// TIA Portal project "消毒机" (V15.1) (continued)
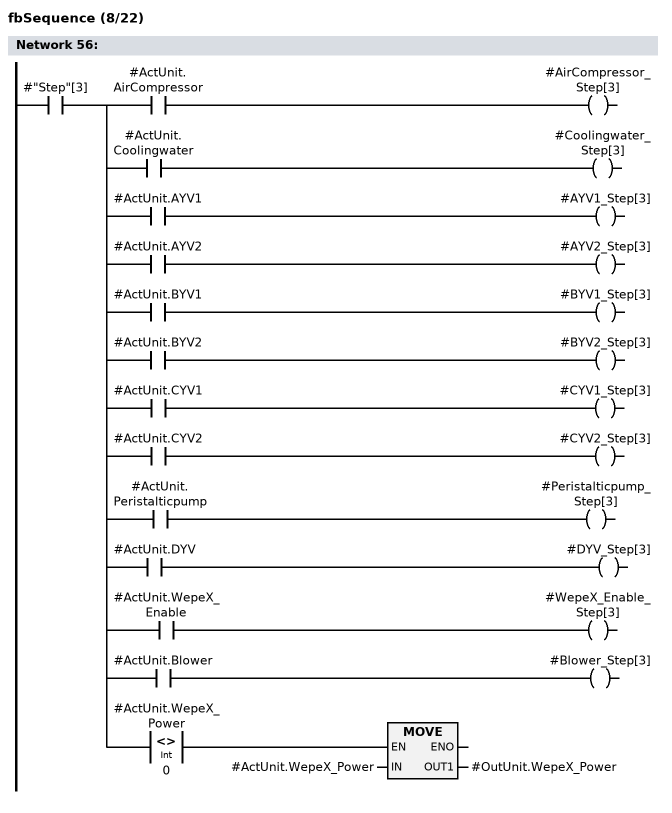
   RUNG wire#powerrail
      Contact( #"Step"[3] )
      wire#w1
      Contact( #ActUnit.AirCompressor )
      Coil( #AirCompressor_Step[3] )
   END_RUNG
   RUNG wire#w1
      Contact( #ActUnit.Coolingwater )
      Coil( #Coolingwater_Step[3] )
   END_RUNG
   RUNG wire#w1
      Contact( #ActUnit.AYV1 )
      Coil( #AYV1_Step[3] )
   END_RUNG
   RUNG wire#w1
      Contact( #ActUnit.AYV2 )
      Coil( #AYV2_Step[3] )
   END_RUNG
   RUNG wire#w1
      Contact( #ActUnit.BYV1 )
      Coil( #BYV1_Step[3] )
   END_RUNG
   RUNG wire#w1
      Contact( #ActUnit.BYV2 )
      Coil( #BYV2_Step[3] )
   END_RUNG
   RUNG wire#w1
      Contact( #ActUnit.CYV1 )
      Coil( #CYV1_Step[3] )
   END_RUNG
   RUNG wire#w1
      Contact( #ActUnit.CYV2 )
      Coil( #CYV2_Step[3] )
   END_RUNG
   RUNG wire#w1
      Contact( #ActUnit.Peristalticpump )
      Coil( #Peristalticpump_Step[3] )
   END_RUNG
   RUNG wire#w1
      Contact( #ActUnit.DYV )
      Coil( #DYV_Step[3] )
   END_RUNG
   RUNG wire#w1
      Contact( #ActUnit.WepeX_Enable )
      Coil( #WepeX_Enable_Step[3] )
   END_RUNG
   RUNG wire#w1
      Contact( #ActUnit.Blower )
      Coil( #Blower_Step[3] )
   END_RUNG
   RUNG wire#w1
      { S7_Templates := "SrcType := Int" } NE_Contact(in1 := #ActUnit.WepeX_Power, in2 := 0)
      Move(in := #ActUnit.WepeX_Power, out1 => #OutUnit.WepeX_Power)
   END_RUNG
   // the same network as SCL:
   #AirCompressor_Step[3] := #"Step"[3] AND #ActUnit.AirCompressor;
   #Coolingwater_Step[3] := #"Step"[3] AND #ActUnit.Coolingwater;
   #AYV1_Step[3] := #"Step"[3] AND #ActUnit.AYV1;
   #AYV2_Step[3] := #"Step"[3] AND #ActUnit.AYV2;
   #BYV1_Step[3] := #"Step"[3] AND #ActUnit.BYV1;
   #BYV2_Step[3] := #"Step"[3] AND #ActUnit.BYV2;
   #CYV1_Step[3] := #"Step"[3] AND #ActUnit.CYV1;
   #CYV2_Step[3] := #"Step"[3] AND #ActUnit.CYV2;
   #Peristalticpump_Step[3] := #"Step"[3] AND #ActUnit.Peristalticpump;
   #DYV_Step[3] := #"Step"[3] AND #ActUnit.DYV;
   #WepeX_Enable_Step[3] := #"Step"[3] AND #ActUnit.WepeX_Enable;
   #Blower_Step[3] := #"Step"[3] AND #ActUnit.Blower;
   IF #"Step"[3] AND (#ActUnit.WepeX_Power <> 0) THEN #OutUnit.WepeX_Power := #ActUnit.WepeX_Power; END_IF;
END_REGION

REGION Network 57
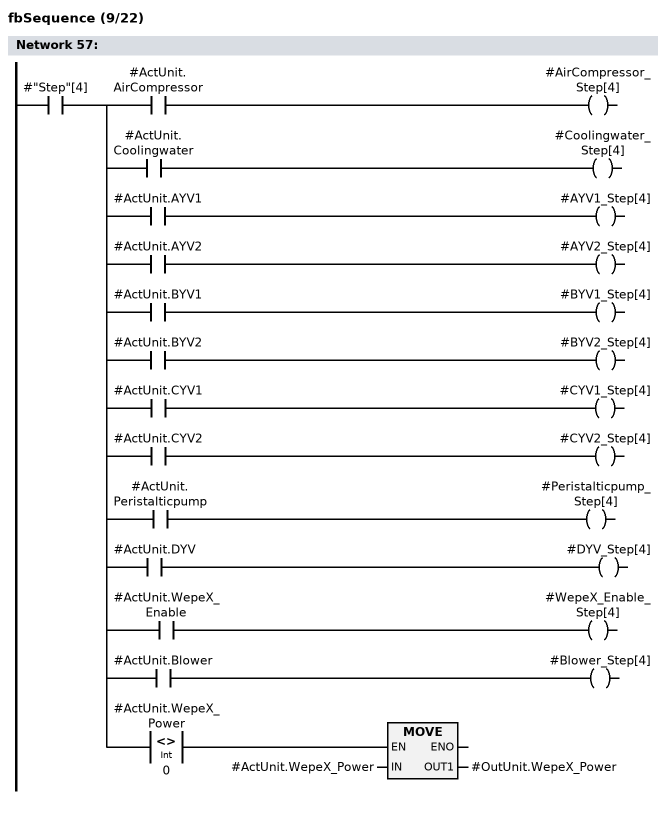
   RUNG wire#powerrail
      Contact( #"Step"[4] )
      wire#w1
      Contact( #ActUnit.AirCompressor )
      Coil( #AirCompressor_Step[4] )
   END_RUNG
   RUNG wire#w1
      Contact( #ActUnit.Coolingwater )
      Coil( #Coolingwater_Step[4] )
   END_RUNG
   RUNG wire#w1
      Contact( #ActUnit.AYV1 )
      Coil( #AYV1_Step[4] )
   END_RUNG
   RUNG wire#w1
      Contact( #ActUnit.AYV2 )
      Coil( #AYV2_Step[4] )
   END_RUNG
   RUNG wire#w1
      Contact( #ActUnit.BYV1 )
      Coil( #BYV1_Step[4] )
   END_RUNG
   RUNG wire#w1
      Contact( #ActUnit.BYV2 )
      Coil( #BYV2_Step[4] )
   END_RUNG
   RUNG wire#w1
      Contact( #ActUnit.CYV1 )
      Coil( #CYV1_Step[4] )
   END_RUNG
   RUNG wire#w1
      Contact( #ActUnit.CYV2 )
      Coil( #CYV2_Step[4] )
   END_RUNG
   RUNG wire#w1
      Contact( #ActUnit.Peristalticpump )
      Coil( #Peristalticpump_Step[4] )
   END_RUNG
   RUNG wire#w1
      Contact( #ActUnit.DYV )
      Coil( #DYV_Step[4] )
   END_RUNG
   RUNG wire#w1
      Contact( #ActUnit.WepeX_Enable )
      Coil( #WepeX_Enable_Step[4] )
   END_RUNG
   RUNG wire#w1
      Contact( #ActUnit.Blower )
      Coil( #Blower_Step[4] )
   END_RUNG
   RUNG wire#w1
      { S7_Templates := "SrcType := Int" } NE_Contact(in1 := #ActUnit.WepeX_Power, in2 := 0)
      Move(in := #ActUnit.WepeX_Power, out1 => #OutUnit.WepeX_Power)
   END_RUNG
   // the same network as SCL:
   #AirCompressor_Step[4] := #"Step"[4] AND #ActUnit.AirCompressor;
   #Coolingwater_Step[4] := #"Step"[4] AND #ActUnit.Coolingwater;
   #AYV1_Step[4] := #"Step"[4] AND #ActUnit.AYV1;
   #AYV2_Step[4] := #"Step"[4] AND #ActUnit.AYV2;
   #BYV1_Step[4] := #"Step"[4] AND #ActUnit.BYV1;
   #BYV2_Step[4] := #"Step"[4] AND #ActUnit.BYV2;
   #CYV1_Step[4] := #"Step"[4] AND #ActUnit.CYV1;
   #CYV2_Step[4] := #"Step"[4] AND #ActUnit.CYV2;
   #Peristalticpump_Step[4] := #"Step"[4] AND #ActUnit.Peristalticpump;
   #DYV_Step[4] := #"Step"[4] AND #ActUnit.DYV;
   #WepeX_Enable_Step[4] := #"Step"[4] AND #ActUnit.WepeX_Enable;
   #Blower_Step[4] := #"Step"[4] AND #ActUnit.Blower;
   IF #"Step"[4] AND (#ActUnit.WepeX_Power <> 0) THEN #OutUnit.WepeX_Power := #ActUnit.WepeX_Power; END_IF;
END_REGION

REGION Network 58
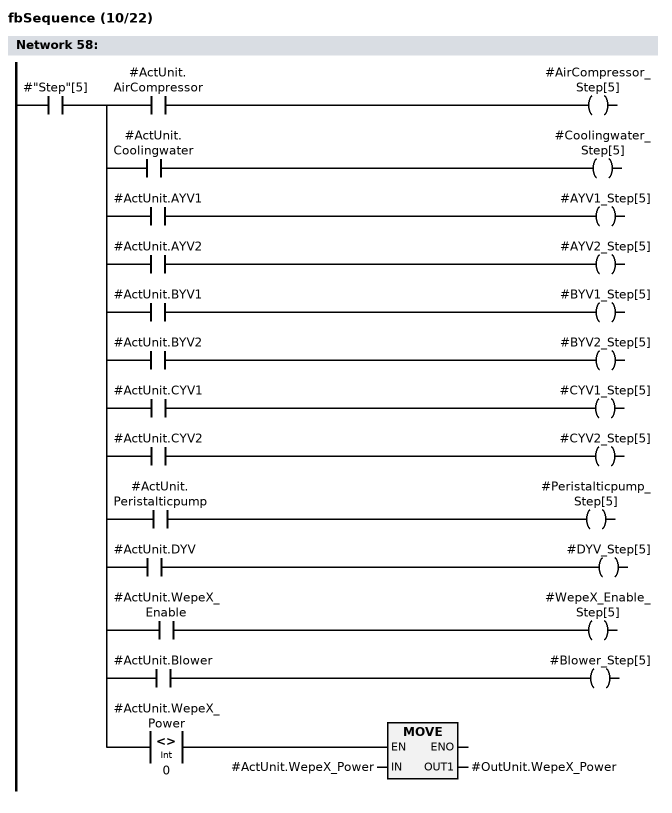
   RUNG wire#powerrail
      Contact( #"Step"[5] )
      wire#w1
      Contact( #ActUnit.AirCompressor )
      Coil( #AirCompressor_Step[5] )
   END_RUNG
   RUNG wire#w1
      Contact( #ActUnit.Coolingwater )
      Coil( #Coolingwater_Step[5] )
   END_RUNG
   RUNG wire#w1
      Contact( #ActUnit.AYV1 )
      Coil( #AYV1_Step[5] )
   END_RUNG
   RUNG wire#w1
      Contact( #ActUnit.AYV2 )
      Coil( #AYV2_Step[5] )
   END_RUNG
   RUNG wire#w1
      Contact( #ActUnit.BYV1 )
      Coil( #BYV1_Step[5] )
   END_RUNG
   RUNG wire#w1
      Contact( #ActUnit.BYV2 )
      Coil( #BYV2_Step[5] )
   END_RUNG
   RUNG wire#w1
      Contact( #ActUnit.CYV1 )
      Coil( #CYV1_Step[5] )
   END_RUNG
   RUNG wire#w1
      Contact( #ActUnit.CYV2 )
      Coil( #CYV2_Step[5] )
   END_RUNG
   RUNG wire#w1
      Contact( #ActUnit.Peristalticpump )
      Coil( #Peristalticpump_Step[5] )
   END_RUNG
   RUNG wire#w1
      Contact( #ActUnit.DYV )
      Coil( #DYV_Step[5] )
   END_RUNG
   RUNG wire#w1
      Contact( #ActUnit.WepeX_Enable )
      Coil( #WepeX_Enable_Step[5] )
   END_RUNG
   RUNG wire#w1
      Contact( #ActUnit.Blower )
      Coil( #Blower_Step[5] )
   END_RUNG
   RUNG wire#w1
      { S7_Templates := "SrcType := Int" } NE_Contact(in1 := #ActUnit.WepeX_Power, in2 := 0)
      Move(in := #ActUnit.WepeX_Power, out1 => #OutUnit.WepeX_Power)
   END_RUNG
   // the same network as SCL:
   #AirCompressor_Step[5] := #"Step"[5] AND #ActUnit.AirCompressor;
   #Coolingwater_Step[5] := #"Step"[5] AND #ActUnit.Coolingwater;
   #AYV1_Step[5] := #"Step"[5] AND #ActUnit.AYV1;
   #AYV2_Step[5] := #"Step"[5] AND #ActUnit.AYV2;
   #BYV1_Step[5] := #"Step"[5] AND #ActUnit.BYV1;
   #BYV2_Step[5] := #"Step"[5] AND #ActUnit.BYV2;
   #CYV1_Step[5] := #"Step"[5] AND #ActUnit.CYV1;
   #CYV2_Step[5] := #"Step"[5] AND #ActUnit.CYV2;
   #Peristalticpump_Step[5] := #"Step"[5] AND #ActUnit.Peristalticpump;
   #DYV_Step[5] := #"Step"[5] AND #ActUnit.DYV;
   #WepeX_Enable_Step[5] := #"Step"[5] AND #ActUnit.WepeX_Enable;
   #Blower_Step[5] := #"Step"[5] AND #ActUnit.Blower;
   IF #"Step"[5] AND (#ActUnit.WepeX_Power <> 0) THEN #OutUnit.WepeX_Power := #ActUnit.WepeX_Power; END_IF;
END_REGION

REGION Network 59
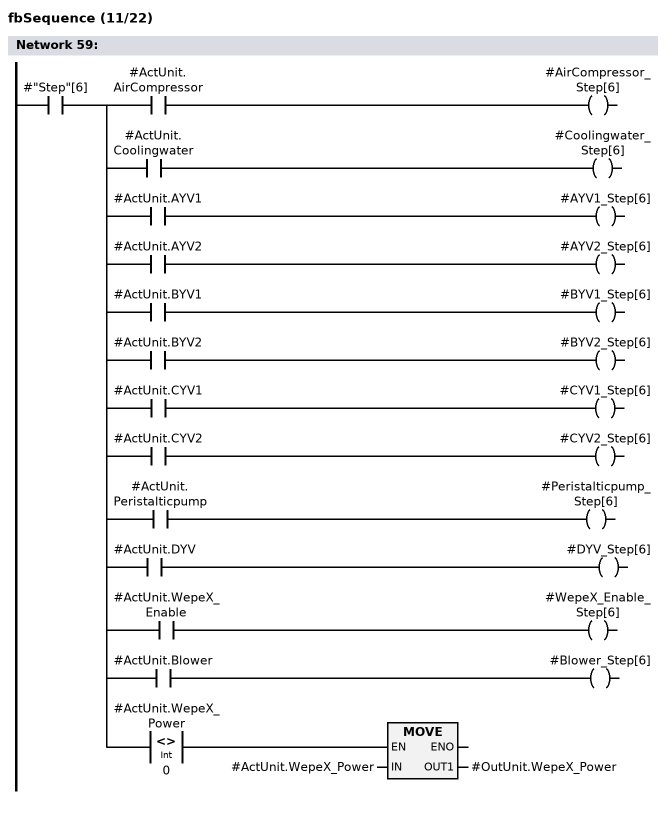
   RUNG wire#powerrail
      Contact( #"Step"[6] )
      wire#w1
      Contact( #ActUnit.AirCompressor )
      Coil( #AirCompressor_Step[6] )
   END_RUNG
   RUNG wire#w1
      Contact( #ActUnit.Coolingwater )
      Coil( #Coolingwater_Step[6] )
   END_RUNG
   RUNG wire#w1
      Contact( #ActUnit.AYV1 )
      Coil( #AYV1_Step[6] )
   END_RUNG
   RUNG wire#w1
      Contact( #ActUnit.AYV2 )
      Coil( #AYV2_Step[6] )
   END_RUNG
   RUNG wire#w1
      Contact( #ActUnit.BYV1 )
      Coil( #BYV1_Step[6] )
   END_RUNG
   RUNG wire#w1
      Contact( #ActUnit.BYV2 )
      Coil( #BYV2_Step[6] )
   END_RUNG
   RUNG wire#w1
      Contact( #ActUnit.CYV1 )
      Coil( #CYV1_Step[6] )
   END_RUNG
   RUNG wire#w1
      Contact( #ActUnit.CYV2 )
      Coil( #CYV2_Step[6] )
   END_RUNG
   RUNG wire#w1
      Contact( #ActUnit.Peristalticpump )
      Coil( #Peristalticpump_Step[6] )
   END_RUNG
   RUNG wire#w1
      Contact( #ActUnit.DYV )
      Coil( #DYV_Step[6] )
   END_RUNG
   RUNG wire#w1
      Contact( #ActUnit.WepeX_Enable )
      Coil( #WepeX_Enable_Step[6] )
   END_RUNG
   RUNG wire#w1
      Contact( #ActUnit.Blower )
      Coil( #Blower_Step[6] )
   END_RUNG
   RUNG wire#w1
      { S7_Templates := "SrcType := Int" } NE_Contact(in1 := #ActUnit.WepeX_Power, in2 := 0)
      Move(in := #ActUnit.WepeX_Power, out1 => #OutUnit.WepeX_Power)
   END_RUNG
   // the same network as SCL:
   #AirCompressor_Step[6] := #"Step"[6] AND #ActUnit.AirCompressor;
   #Coolingwater_Step[6] := #"Step"[6] AND #ActUnit.Coolingwater;
   #AYV1_Step[6] := #"Step"[6] AND #ActUnit.AYV1;
   #AYV2_Step[6] := #"Step"[6] AND #ActUnit.AYV2;
   #BYV1_Step[6] := #"Step"[6] AND #ActUnit.BYV1;
   #BYV2_Step[6] := #"Step"[6] AND #ActUnit.BYV2;
   #CYV1_Step[6] := #"Step"[6] AND #ActUnit.CYV1;
   #CYV2_Step[6] := #"Step"[6] AND #ActUnit.CYV2;
   #Peristalticpump_Step[6] := #"Step"[6] AND #ActUnit.Peristalticpump;
   #DYV_Step[6] := #"Step"[6] AND #ActUnit.DYV;
   #WepeX_Enable_Step[6] := #"Step"[6] AND #ActUnit.WepeX_Enable;
   #Blower_Step[6] := #"Step"[6] AND #ActUnit.Blower;
   IF #"Step"[6] AND (#ActUnit.WepeX_Power <> 0) THEN #OutUnit.WepeX_Power := #ActUnit.WepeX_Power; END_IF;
END_REGION

REGION Network 60
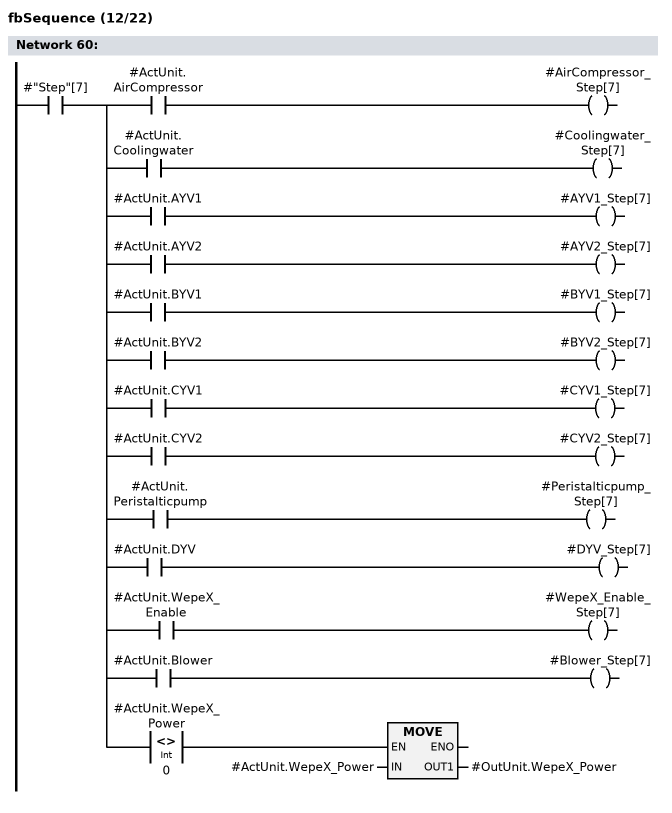
   RUNG wire#powerrail
      Contact( #"Step"[7] )
      wire#w1
      Contact( #ActUnit.AirCompressor )
      Coil( #AirCompressor_Step[7] )
   END_RUNG
   RUNG wire#w1
      Contact( #ActUnit.Coolingwater )
      Coil( #Coolingwater_Step[7] )
   END_RUNG
   RUNG wire#w1
      Contact( #ActUnit.AYV1 )
      Coil( #AYV1_Step[7] )
   END_RUNG
   RUNG wire#w1
      Contact( #ActUnit.AYV2 )
      Coil( #AYV2_Step[7] )
   END_RUNG
   RUNG wire#w1
      Contact( #ActUnit.BYV1 )
      Coil( #BYV1_Step[7] )
   END_RUNG
   RUNG wire#w1
      Contact( #ActUnit.BYV2 )
      Coil( #BYV2_Step[7] )
   END_RUNG
   RUNG wire#w1
      Contact( #ActUnit.CYV1 )
      Coil( #CYV1_Step[7] )
   END_RUNG
   RUNG wire#w1
      Contact( #ActUnit.CYV2 )
      Coil( #CYV2_Step[7] )
   END_RUNG
   RUNG wire#w1
      Contact( #ActUnit.Peristalticpump )
      Coil( #Peristalticpump_Step[7] )
   END_RUNG
   RUNG wire#w1
      Contact( #ActUnit.DYV )
      Coil( #DYV_Step[7] )
   END_RUNG
   RUNG wire#w1
      Contact( #ActUnit.WepeX_Enable )
      Coil( #WepeX_Enable_Step[7] )
   END_RUNG
   RUNG wire#w1
      Contact( #ActUnit.Blower )
      Coil( #Blower_Step[7] )
   END_RUNG
   RUNG wire#w1
      { S7_Templates := "SrcType := Int" } NE_Contact(in1 := #ActUnit.WepeX_Power, in2 := 0)
      Move(in := #ActUnit.WepeX_Power, out1 => #OutUnit.WepeX_Power)
   END_RUNG
   // the same network as SCL:
   #AirCompressor_Step[7] := #"Step"[7] AND #ActUnit.AirCompressor;
   #Coolingwater_Step[7] := #"Step"[7] AND #ActUnit.Coolingwater;
   #AYV1_Step[7] := #"Step"[7] AND #ActUnit.AYV1;
   #AYV2_Step[7] := #"Step"[7] AND #ActUnit.AYV2;
   #BYV1_Step[7] := #"Step"[7] AND #ActUnit.BYV1;
   #BYV2_Step[7] := #"Step"[7] AND #ActUnit.BYV2;
   #CYV1_Step[7] := #"Step"[7] AND #ActUnit.CYV1;
   #CYV2_Step[7] := #"Step"[7] AND #ActUnit.CYV2;
   #Peristalticpump_Step[7] := #"Step"[7] AND #ActUnit.Peristalticpump;
   #DYV_Step[7] := #"Step"[7] AND #ActUnit.DYV;
   #WepeX_Enable_Step[7] := #"Step"[7] AND #ActUnit.WepeX_Enable;
   #Blower_Step[7] := #"Step"[7] AND #ActUnit.Blower;
   IF #"Step"[7] AND (#ActUnit.WepeX_Power <> 0) THEN #OutUnit.WepeX_Power := #ActUnit.WepeX_Power; END_IF;
END_REGION

REGION Network 61
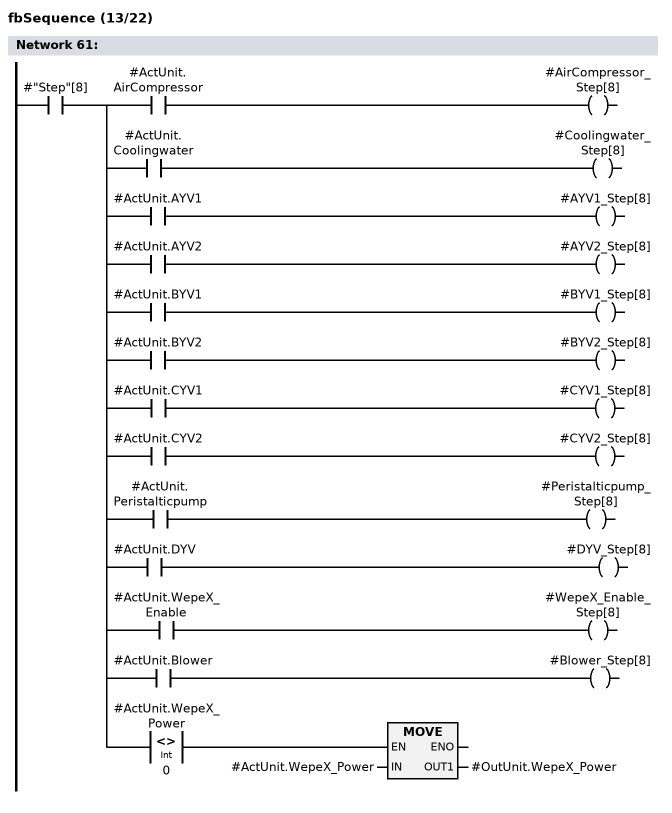
   RUNG wire#powerrail
      Contact( #"Step"[8] )
      wire#w1
      Contact( #ActUnit.AirCompressor )
      Coil( #AirCompressor_Step[8] )
   END_RUNG
   RUNG wire#w1
      Contact( #ActUnit.Coolingwater )
      Coil( #Coolingwater_Step[8] )
   END_RUNG
   RUNG wire#w1
      Contact( #ActUnit.AYV1 )
      Coil( #AYV1_Step[8] )
   END_RUNG
   RUNG wire#w1
      Contact( #ActUnit.AYV2 )
      Coil( #AYV2_Step[8] )
   END_RUNG
   RUNG wire#w1
      Contact( #ActUnit.BYV1 )
      Coil( #BYV1_Step[8] )
   END_RUNG
   RUNG wire#w1
      Contact( #ActUnit.BYV2 )
      Coil( #BYV2_Step[8] )
   END_RUNG
   RUNG wire#w1
      Contact( #ActUnit.CYV1 )
      Coil( #CYV1_Step[8] )
   END_RUNG
   RUNG wire#w1
      Contact( #ActUnit.CYV2 )
      Coil( #CYV2_Step[8] )
   END_RUNG
   RUNG wire#w1
      Contact( #ActUnit.Peristalticpump )
      Coil( #Peristalticpump_Step[8] )
   END_RUNG
   RUNG wire#w1
      Contact( #ActUnit.DYV )
      Coil( #DYV_Step[8] )
   END_RUNG
   RUNG wire#w1
      Contact( #ActUnit.WepeX_Enable )
      Coil( #WepeX_Enable_Step[8] )
   END_RUNG
   RUNG wire#w1
      Contact( #ActUnit.Blower )
      Coil( #Blower_Step[8] )
   END_RUNG
   RUNG wire#w1
      { S7_Templates := "SrcType := Int" } NE_Contact(in1 := #ActUnit.WepeX_Power, in2 := 0)
      Move(in := #ActUnit.WepeX_Power, out1 => #OutUnit.WepeX_Power)
   END_RUNG
   // the same network as SCL:
   #AirCompressor_Step[8] := #"Step"[8] AND #ActUnit.AirCompressor;
   #Coolingwater_Step[8] := #"Step"[8] AND #ActUnit.Coolingwater;
   #AYV1_Step[8] := #"Step"[8] AND #ActUnit.AYV1;
   #AYV2_Step[8] := #"Step"[8] AND #ActUnit.AYV2;
   #BYV1_Step[8] := #"Step"[8] AND #ActUnit.BYV1;
   #BYV2_Step[8] := #"Step"[8] AND #ActUnit.BYV2;
   #CYV1_Step[8] := #"Step"[8] AND #ActUnit.CYV1;
   #CYV2_Step[8] := #"Step"[8] AND #ActUnit.CYV2;
   #Peristalticpump_Step[8] := #"Step"[8] AND #ActUnit.Peristalticpump;
   #DYV_Step[8] := #"Step"[8] AND #ActUnit.DYV;
   #WepeX_Enable_Step[8] := #"Step"[8] AND #ActUnit.WepeX_Enable;
   #Blower_Step[8] := #"Step"[8] AND #ActUnit.Blower;
   IF #"Step"[8] AND (#ActUnit.WepeX_Power <> 0) THEN #OutUnit.WepeX_Power := #ActUnit.WepeX_Power; END_IF;
END_REGION

REGION Network 62
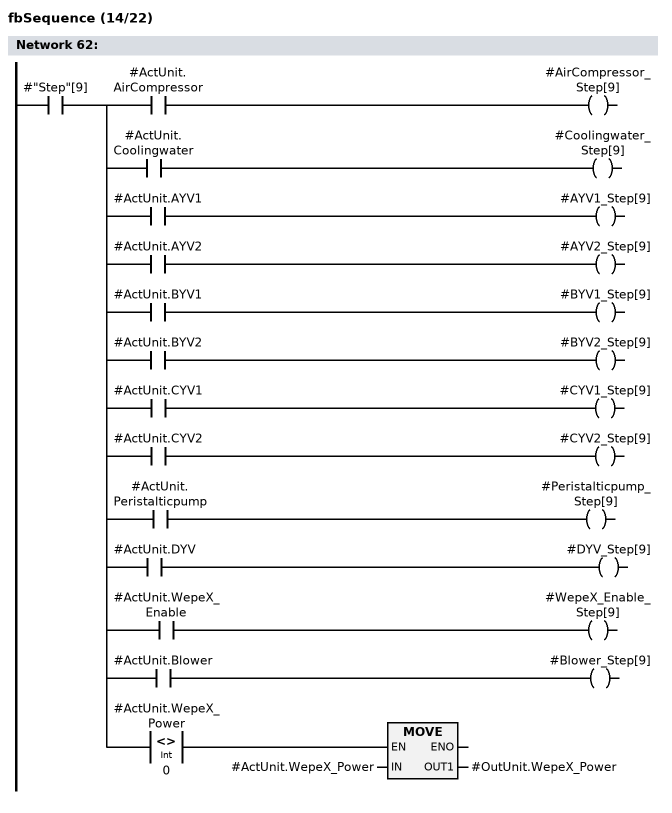
   RUNG wire#powerrail
      Contact( #"Step"[9] )
      wire#w1
      Contact( #ActUnit.AirCompressor )
      Coil( #AirCompressor_Step[9] )
   END_RUNG
   RUNG wire#w1
      Contact( #ActUnit.Coolingwater )
      Coil( #Coolingwater_Step[9] )
   END_RUNG
   RUNG wire#w1
      Contact( #ActUnit.AYV1 )
      Coil( #AYV1_Step[9] )
   END_RUNG
   RUNG wire#w1
      Contact( #ActUnit.AYV2 )
      Coil( #AYV2_Step[9] )
   END_RUNG
   RUNG wire#w1
      Contact( #ActUnit.BYV1 )
      Coil( #BYV1_Step[9] )
   END_RUNG
   RUNG wire#w1
      Contact( #ActUnit.BYV2 )
      Coil( #BYV2_Step[9] )
   END_RUNG
   RUNG wire#w1
      Contact( #ActUnit.CYV1 )
      Coil( #CYV1_Step[9] )
   END_RUNG
   RUNG wire#w1
      Contact( #ActUnit.CYV2 )
      Coil( #CYV2_Step[9] )
   END_RUNG
   RUNG wire#w1
      Contact( #ActUnit.Peristalticpump )
      Coil( #Peristalticpump_Step[9] )
   END_RUNG
   RUNG wire#w1
      Contact( #ActUnit.DYV )
      Coil( #DYV_Step[9] )
   END_RUNG
   RUNG wire#w1
      Contact( #ActUnit.WepeX_Enable )
      Coil( #WepeX_Enable_Step[9] )
   END_RUNG
   RUNG wire#w1
      Contact( #ActUnit.Blower )
      Coil( #Blower_Step[9] )
   END_RUNG
   RUNG wire#w1
      { S7_Templates := "SrcType := Int" } NE_Contact(in1 := #ActUnit.WepeX_Power, in2 := 0)
      Move(in := #ActUnit.WepeX_Power, out1 => #OutUnit.WepeX_Power)
   END_RUNG
   // the same network as SCL:
   #AirCompressor_Step[9] := #"Step"[9] AND #ActUnit.AirCompressor;
   #Coolingwater_Step[9] := #"Step"[9] AND #ActUnit.Coolingwater;
   #AYV1_Step[9] := #"Step"[9] AND #ActUnit.AYV1;
   #AYV2_Step[9] := #"Step"[9] AND #ActUnit.AYV2;
   #BYV1_Step[9] := #"Step"[9] AND #ActUnit.BYV1;
   #BYV2_Step[9] := #"Step"[9] AND #ActUnit.BYV2;
   #CYV1_Step[9] := #"Step"[9] AND #ActUnit.CYV1;
   #CYV2_Step[9] := #"Step"[9] AND #ActUnit.CYV2;
   #Peristalticpump_Step[9] := #"Step"[9] AND #ActUnit.Peristalticpump;
   #DYV_Step[9] := #"Step"[9] AND #ActUnit.DYV;
   #WepeX_Enable_Step[9] := #"Step"[9] AND #ActUnit.WepeX_Enable;
   #Blower_Step[9] := #"Step"[9] AND #ActUnit.Blower;
   IF #"Step"[9] AND (#ActUnit.WepeX_Power <> 0) THEN #OutUnit.WepeX_Power := #ActUnit.WepeX_Power; END_IF;
END_REGION

REGION Network 63
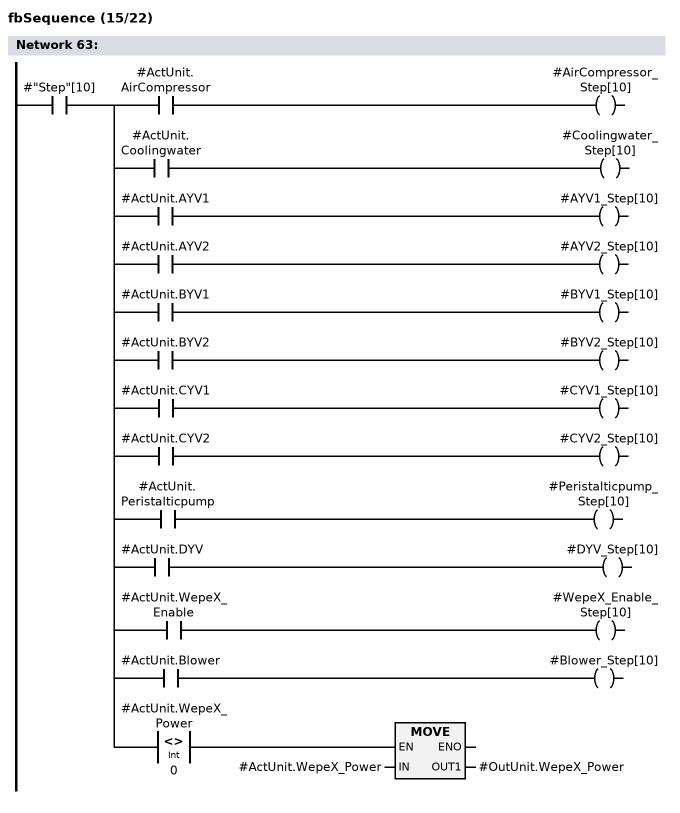
   RUNG wire#powerrail
      Contact( #"Step"[10] )
      wire#w1
      Contact( #ActUnit.AirCompressor )
      Coil( #AirCompressor_Step[10] )
   END_RUNG
   RUNG wire#w1
      Contact( #ActUnit.Coolingwater )
      Coil( #Coolingwater_Step[10] )
   END_RUNG
   RUNG wire#w1
      Contact( #ActUnit.AYV1 )
      Coil( #AYV1_Step[10] )
   END_RUNG
   RUNG wire#w1
      Contact( #ActUnit.AYV2 )
      Coil( #AYV2_Step[10] )
   END_RUNG
   RUNG wire#w1
      Contact( #ActUnit.BYV1 )
      Coil( #BYV1_Step[10] )
   END_RUNG
   RUNG wire#w1
      Contact( #ActUnit.BYV2 )
      Coil( #BYV2_Step[10] )
   END_RUNG
   RUNG wire#w1
      Contact( #ActUnit.CYV1 )
      Coil( #CYV1_Step[10] )
   END_RUNG
   RUNG wire#w1
      Contact( #ActUnit.CYV2 )
      Coil( #CYV2_Step[10] )
   END_RUNG
   RUNG wire#w1
      Contact( #ActUnit.Peristalticpump )
      Coil( #Peristalticpump_Step[10] )
   END_RUNG
   RUNG wire#w1
      Contact( #ActUnit.DYV )
      Coil( #DYV_Step[10] )
   END_RUNG
   RUNG wire#w1
      Contact( #ActUnit.WepeX_Enable )
      Coil( #WepeX_Enable_Step[10] )
   END_RUNG
   RUNG wire#w1
      Contact( #ActUnit.Blower )
      Coil( #Blower_Step[10] )
   END_RUNG
   RUNG wire#w1
      { S7_Templates := "SrcType := Int" } NE_Contact(in1 := #ActUnit.WepeX_Power, in2 := 0)
      Move(in := #ActUnit.WepeX_Power, out1 => #OutUnit.WepeX_Power)
   END_RUNG
   // the same network as SCL:
   #AirCompressor_Step[10] := #"Step"[10] AND #ActUnit.AirCompressor;
   #Coolingwater_Step[10] := #"Step"[10] AND #ActUnit.Coolingwater;
   #AYV1_Step[10] := #"Step"[10] AND #ActUnit.AYV1;
   #AYV2_Step[10] := #"Step"[10] AND #ActUnit.AYV2;
   #BYV1_Step[10] := #"Step"[10] AND #ActUnit.BYV1;
   #BYV2_Step[10] := #"Step"[10] AND #ActUnit.BYV2;
   #CYV1_Step[10] := #"Step"[10] AND #ActUnit.CYV1;
   #CYV2_Step[10] := #"Step"[10] AND #ActUnit.CYV2;
   #Peristalticpump_Step[10] := #"Step"[10] AND #ActUnit.Peristalticpump;
   #DYV_Step[10] := #"Step"[10] AND #ActUnit.DYV;
   #WepeX_Enable_Step[10] := #"Step"[10] AND #ActUnit.WepeX_Enable;
   #Blower_Step[10] := #"Step"[10] AND #ActUnit.Blower;
   IF #"Step"[10] AND (#ActUnit.WepeX_Power <> 0) THEN #OutUnit.WepeX_Power := #ActUnit.WepeX_Power; END_IF;
END_REGION

REGION Network 64
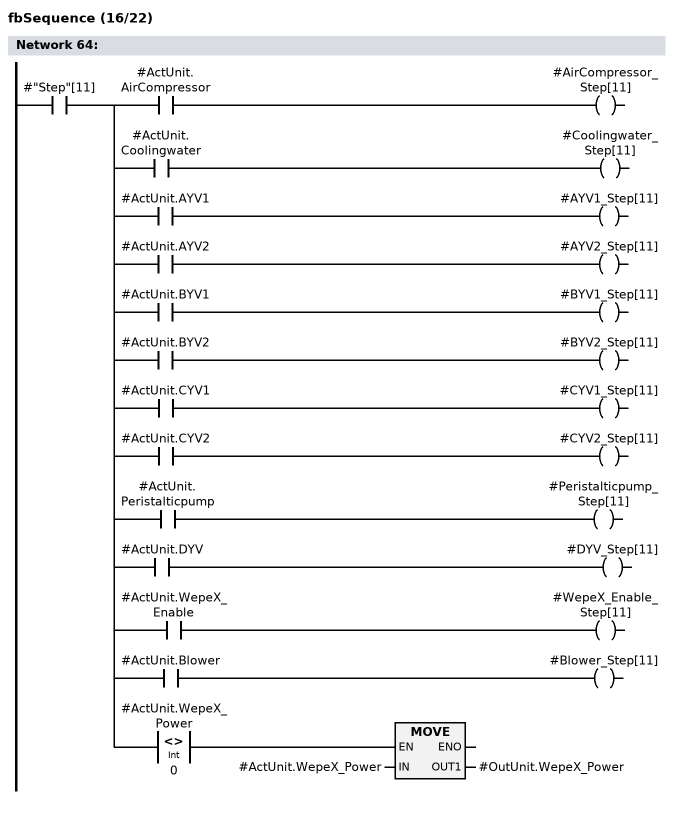
   RUNG wire#powerrail
      Contact( #"Step"[11] )
      wire#w1
      Contact( #ActUnit.AirCompressor )
      Coil( #AirCompressor_Step[11] )
   END_RUNG
   RUNG wire#w1
      Contact( #ActUnit.Coolingwater )
      Coil( #Coolingwater_Step[11] )
   END_RUNG
   RUNG wire#w1
      Contact( #ActUnit.AYV1 )
      Coil( #AYV1_Step[11] )
   END_RUNG
   RUNG wire#w1
      Contact( #ActUnit.AYV2 )
      Coil( #AYV2_Step[11] )
   END_RUNG
   RUNG wire#w1
      Contact( #ActUnit.BYV1 )
      Coil( #BYV1_Step[11] )
   END_RUNG
   RUNG wire#w1
      Contact( #ActUnit.BYV2 )
      Coil( #BYV2_Step[11] )
   END_RUNG
   RUNG wire#w1
      Contact( #ActUnit.CYV1 )
      Coil( #CYV1_Step[11] )
   END_RUNG
   RUNG wire#w1
      Contact( #ActUnit.CYV2 )
      Coil( #CYV2_Step[11] )
   END_RUNG
   RUNG wire#w1
      Contact( #ActUnit.Peristalticpump )
      Coil( #Peristalticpump_Step[11] )
   END_RUNG
   RUNG wire#w1
      Contact( #ActUnit.DYV )
      Coil( #DYV_Step[11] )
   END_RUNG
   RUNG wire#w1
      Contact( #ActUnit.WepeX_Enable )
      Coil( #WepeX_Enable_Step[11] )
   END_RUNG
   RUNG wire#w1
      Contact( #ActUnit.Blower )
      Coil( #Blower_Step[11] )
   END_RUNG
   RUNG wire#w1
      { S7_Templates := "SrcType := Int" } NE_Contact(in1 := #ActUnit.WepeX_Power, in2 := 0)
      Move(in := #ActUnit.WepeX_Power, out1 => #OutUnit.WepeX_Power)
   END_RUNG
   // the same network as SCL:
   #AirCompressor_Step[11] := #"Step"[11] AND #ActUnit.AirCompressor;
   #Coolingwater_Step[11] := #"Step"[11] AND #ActUnit.Coolingwater;
   #AYV1_Step[11] := #"Step"[11] AND #ActUnit.AYV1;
   #AYV2_Step[11] := #"Step"[11] AND #ActUnit.AYV2;
   #BYV1_Step[11] := #"Step"[11] AND #ActUnit.BYV1;
   #BYV2_Step[11] := #"Step"[11] AND #ActUnit.BYV2;
   #CYV1_Step[11] := #"Step"[11] AND #ActUnit.CYV1;
   #CYV2_Step[11] := #"Step"[11] AND #ActUnit.CYV2;
   #Peristalticpump_Step[11] := #"Step"[11] AND #ActUnit.Peristalticpump;
   #DYV_Step[11] := #"Step"[11] AND #ActUnit.DYV;
   #WepeX_Enable_Step[11] := #"Step"[11] AND #ActUnit.WepeX_Enable;
   #Blower_Step[11] := #"Step"[11] AND #ActUnit.Blower;
   IF #"Step"[11] AND (#ActUnit.WepeX_Power <> 0) THEN #OutUnit.WepeX_Power := #ActUnit.WepeX_Power; END_IF;
END_REGION

REGION Network 65
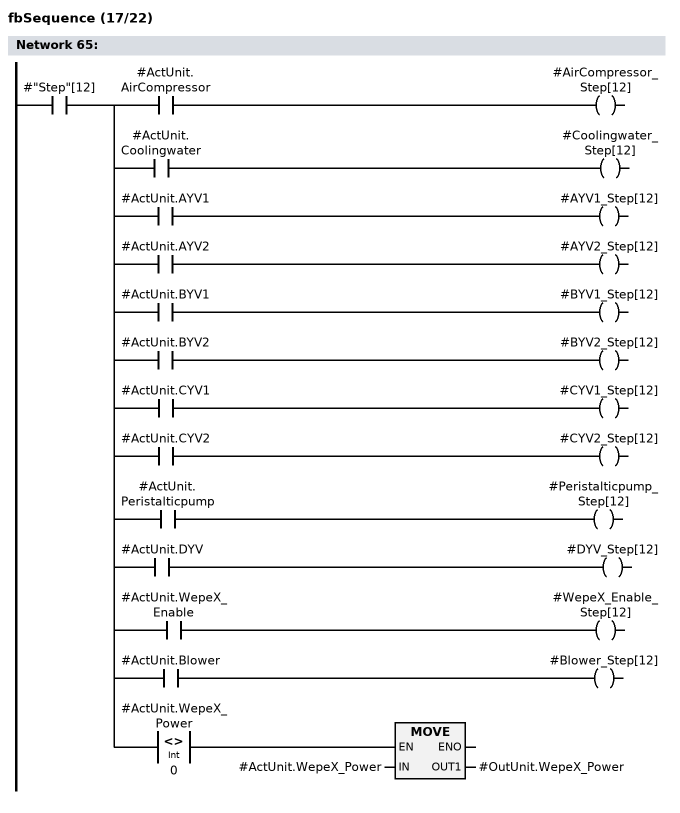
   RUNG wire#powerrail
      Contact( #"Step"[12] )
      wire#w1
      Contact( #ActUnit.AirCompressor )
      Coil( #AirCompressor_Step[12] )
   END_RUNG
   RUNG wire#w1
      Contact( #ActUnit.Coolingwater )
      Coil( #Coolingwater_Step[12] )
   END_RUNG
   RUNG wire#w1
      Contact( #ActUnit.AYV1 )
      Coil( #AYV1_Step[12] )
   END_RUNG
   RUNG wire#w1
      Contact( #ActUnit.AYV2 )
      Coil( #AYV2_Step[12] )
   END_RUNG
   RUNG wire#w1
      Contact( #ActUnit.BYV1 )
      Coil( #BYV1_Step[12] )
   END_RUNG
   RUNG wire#w1
      Contact( #ActUnit.BYV2 )
      Coil( #BYV2_Step[12] )
   END_RUNG
   RUNG wire#w1
      Contact( #ActUnit.CYV1 )
      Coil( #CYV1_Step[12] )
   END_RUNG
   RUNG wire#w1
      Contact( #ActUnit.CYV2 )
      Coil( #CYV2_Step[12] )
   END_RUNG
   RUNG wire#w1
      Contact( #ActUnit.Peristalticpump )
      Coil( #Peristalticpump_Step[12] )
   END_RUNG
   RUNG wire#w1
      Contact( #ActUnit.DYV )
      Coil( #DYV_Step[12] )
   END_RUNG
   RUNG wire#w1
      Contact( #ActUnit.WepeX_Enable )
      Coil( #WepeX_Enable_Step[12] )
   END_RUNG
   RUNG wire#w1
      Contact( #ActUnit.Blower )
      Coil( #Blower_Step[12] )
   END_RUNG
   RUNG wire#w1
      { S7_Templates := "SrcType := Int" } NE_Contact(in1 := #ActUnit.WepeX_Power, in2 := 0)
      Move(in := #ActUnit.WepeX_Power, out1 => #OutUnit.WepeX_Power)
   END_RUNG
   // the same network as SCL:
   #AirCompressor_Step[12] := #"Step"[12] AND #ActUnit.AirCompressor;
   #Coolingwater_Step[12] := #"Step"[12] AND #ActUnit.Coolingwater;
   #AYV1_Step[12] := #"Step"[12] AND #ActUnit.AYV1;
   #AYV2_Step[12] := #"Step"[12] AND #ActUnit.AYV2;
   #BYV1_Step[12] := #"Step"[12] AND #ActUnit.BYV1;
   #BYV2_Step[12] := #"Step"[12] AND #ActUnit.BYV2;
   #CYV1_Step[12] := #"Step"[12] AND #ActUnit.CYV1;
   #CYV2_Step[12] := #"Step"[12] AND #ActUnit.CYV2;
   #Peristalticpump_Step[12] := #"Step"[12] AND #ActUnit.Peristalticpump;
   #DYV_Step[12] := #"Step"[12] AND #ActUnit.DYV;
   #WepeX_Enable_Step[12] := #"Step"[12] AND #ActUnit.WepeX_Enable;
   #Blower_Step[12] := #"Step"[12] AND #ActUnit.Blower;
   IF #"Step"[12] AND (#ActUnit.WepeX_Power <> 0) THEN #OutUnit.WepeX_Power := #ActUnit.WepeX_Power; END_IF;
END_REGION

REGION Network 66
